           // ******************************************************************************************************
       100:  // Error state
           IF #ILx2T_Ref.ProChAccessID = #inAccessID THEN
               #ILx2T_Ref.ProChAccessID := 0;   // release access to proccessdata channel
           END_IF;
           #q_xBusy := FALSE;
           #q_xError := TRUE;
           #inState := 110;
           // ******************************************************************************************************
       110:  // finished
           IF NOT #i_xForward AND NOT #i_xBackward THEN
               #q_xError := FALSE;
               #q_xBusy := FALSE;
               #q_xCommandAborted := FALSE;
               #inState := 0;
           END_IF;
           // ******************************************************************************************************
   END_CASE;
END_FUNCTION_BLOCK

FUNCTION_BLOCK "ILx2T_Parameter_Read_Write"   // FB5, SCL
{ S7_Optimized_Access := 'TRUE' }
VERSION : 1.5
   VAR_INPUT
      i_xParameterRead : Bool;   // TRUE = Reading value continuously
      i_xParameterWrite : Bool;   // rising edge = Writing once
      i_woParameterAddress : Word;   // Parameter address (see product manual)
      i_byWriteParameterLength : Byte;   // parameter length in bytes ( 2 or 4 bytes)
      i_diWriteParameterValue : DInt;   // parameter write value
   END_VAR
   VAR_OUTPUT
      q_xReadValueValid : Bool;   // reading value is valid
      q_xWriteDone : Bool;   // writing finished without error
      q_xError : Bool;   // finished with error
      q_xBusy : Bool;   // function is active
      q_diReadParameterValue : DInt;   // reading value
   END_VAR
   VAR_IN_OUT
      ILx2T_Ref : "ILx2T_Ref";   // Axis reference structure
   END_VAR
   VAR
      inState : Int;   // internal state machine
      inAccessID : Int;   // own access ID
      inErrorState : Int;
      dwParaChErrorNo : DWord;   // parameter channe error ID
      xHelperWrite : Bool;
      xHelperRead : Bool;
      TON_Timeout : TON_TIME;
   END_VAR
BEGIN
   // *******************************************************************************
   // Init after Restart
   // *******************************************************************************
   // Check for PLC restart (1st call of this FB)
   IF #inAccessID = 0 THEN
       #ILx2T_Ref.InitAccessID := #ILx2T_Ref.InitAccessID + 1;
       #inAccessID := #ILx2T_Ref.InitAccessID;
   END_IF;

   CASE #inState OF
           // ******************************************************************************************************
       0:  // idle state
           IF #i_xParameterWrite XOR #i_xParameterRead THEN
               #xHelperWrite := #i_xParameterWrite;
               #xHelperRead := #i_xParameterRead;
               #q_xBusy := TRUE;
               #inErrorState := 0;
               #dwParaChErrorNo := 0;
               #inState := #inState + 1;
           ELSE
               #q_xWriteDone := FALSE;
               #q_xError := FALSE;
               #q_xBusy := FALSE;
               #q_xReadValueValid := FALSE;
               #q_diReadParameterValue := 0;
           END_IF;
           // ******************************************************************************************************
       1:  // Check for parameterchannel access
           IF #ILx2T_Ref.ParChAccessID = 0 OR #ILx2T_Ref.ParChAccessID = #inAccessID THEN
               #ILx2T_Ref.ParChAccessID := #inAccessID;   // grab access to parameter channel
               #inState := #inState + 1;
           END_IF;
           // ******************************************************************************************************
       2:// Prepare parameterchannel command
           #TON_Timeout(IN := FALSE,
                        PT := t#1s);
           IF #xHelperRead THEN
               #ILx2T_Ref.x_CommandReadParameter := TRUE;
               #ILx2T_Ref.udi_ModbusAddress_Read := #i_woParameterAddress;
               #inState := #inState + 1;
           ELSIF #xHelperWrite THEN
               #ILx2T_Ref.x_CommandWriteParameter := TRUE;
               #ILx2T_Ref.udi_ModbusAddress_Write := #i_woParameterAddress;
               #ILx2T_Ref.di_ParameterWriteValue := #i_diWriteParameterValue;
               #inState := #inState + 1;
           END_IF;
           // ******************************************************************************************************
       3: // Check for Parameterchannel response
           #TON_Timeout(IN := TRUE,
                        PT := t#1s);
           IF #TON_Timeout.Q THEN
               #TON_Timeout(IN := FALSE,
                            PT := t#1s);
               #q_xError := TRUE;
               #inErrorState := #inState;
               #inState := 100;
               // Read Done    
           ELSIF #xHelperRead AND #ILx2T_Ref.x_StatusReadParameter_OK AND NOT #ILx2T_Ref.x_StatusReadParameter_Error THEN
               #TON_Timeout(IN := FALSE,
                            PT := t#1s);
               #q_diReadParameterValue := #ILx2T_Ref.di_ParameterReadValue;
               #q_xReadValueValid := TRUE;
               #ILx2T_Ref.x_CommandReadParameter := FALSE;
               #ILx2T_Ref.x_StatusReadParameter_OK := FALSE;
               #ILx2T_Ref.udi_ModbusAddress_Read := 0;
               #inState := #inState + 1;
               // Write Done    
           ELSIF #xHelperWrite AND #ILx2T_Ref.x_Status_WriteParameter_OK AND NOT #ILx2T_Ref.x_Status_WriteParameter_Error THEN
               #TON_Timeout(IN := FALSE,
                            PT := t#1s);
               #ILx2T_Ref.di_ParameterWriteValue := 0;
               #q_xWriteDone := TRUE;
               #ILx2T_Ref.x_CommandWriteParameter := FALSE;
               #ILx2T_Ref.x_Status_WriteParameter_OK := FALSE;
               #ILx2T_Ref.udi_ModbusAddress_Write := 0;
               #inState := #inState + 1;
               // Error response Reading
           ELSIF #ILx2T_Ref.x_StatusReadParameter_Error THEN
               #ILx2T_Ref.x_CommandReadParameter := FALSE;
               #ILx2T_Ref.x_StatusReadParameter_Error := FALSE;
               #ILx2T_Ref.udi_ModbusAddress_Read := 0;
               #TON_Timeout(IN := FALSE,
                            PT := t#1s);
               #inErrorState := #inState;
               #inState := 100;
               // Error response Writing
           ELSIF #ILx2T_Ref.x_Status_WriteParameter_Error THEN
               #ILx2T_Ref.x_CommandWriteParameter := FALSE;
               #ILx2T_Ref.x_Status_WriteParameter_Error := FALSE;
               #ILx2T_Ref.udi_ModbusAddress_Write := 0;
               #TON_Timeout(IN := FALSE,
                            PT := t#1s);
               #inErrorState := #inState;
               #inState := 100;
           END_IF;
           // ******************************************************************************************************
       4:  // Check for Parameterchannel in idle state
           #TON_Timeout(IN := TRUE,
                        PT := t#1s);
           IF #TON_Timeout.Q THEN
               #TON_Timeout(IN := FALSE,
                            PT := t#1s);
               #q_xError := TRUE;
               #inErrorState := #inState;
               #inState := 100;
           ELSIF NOT #ILx2T_Ref.x_StatusReadParameter_OK AND NOT #ILx2T_Ref.x_StatusReadParameter_Error
               AND NOT #ILx2T_Ref.x_Status_WriteParameter_OK AND NOT #ILx2T_Ref.x_Status_WriteParameter_Error THEN
               #ILx2T_Ref.ParChAccessID := 0;   // grab access to parameter channel
               #TON_Timeout(IN := FALSE,
                            PT := t#1s);
               IF #xHelperWrite THEN
                   #q_xBusy := FALSE;
                   #inState := 110;
               ELSE
                   #inState := 0;
               END_IF;
           END_IF;
       100:  // Error state
           IF #ILx2T_Ref.ParChAccessID = #inAccessID THEN
               #ILx2T_Ref.ParChAccessID := 0;   // release access to proccessdata channel
           END_IF;
           #q_xBusy := FALSE;
           #q_xError := TRUE;
           #inState := 110;
           // ******************************************************************************************************
       110:  // finished
           IF NOT #i_xParameterWrite AND NOT #i_xParameterRead THEN
               #q_xWriteDone := FALSE;
               #q_xError := FALSE;
               #q_xBusy := FALSE;
               #q_xReadValueValid := FALSE;
               #q_diReadParameterValue := 0;
               #inState := 0;
           END_IF;
           // ******************************************************************************************************
   END_CASE;
END_FUNCTION_BLOCK

FUNCTION_BLOCK "ILx2T_ProfilePosition"   // FB6, SCL
{ S7_Optimized_Access := 'TRUE' }
VERSION : 1.5
   VAR_INPUT
      i_xExecute : Bool;   // rising edge starts a new movement
      i_xAbort : Bool;   // abort active movement
      i_inPTP_Type : Int;   // 1=absolute / 2=additive / 3=relative
      i_diTargetPosition : DInt;   // Target position value
      i_inTargetVelocity : Int;   // Target velocity value
   END_VAR
   VAR_OUTPUT
      q_xDone : Bool;   // Target position reached
      q_xError : Bool;   // finished with error
      q_xCommandAborted : Bool;   // function aborted
      q_xBusy : Bool;   // function is active
   END_VAR
   VAR_IN_OUT
      ILx2T_Ref : "ILx2T_Ref";   // Axis reference structure
   END_VAR
   VAR
      inState : Int;   // internal state machine
      inAccessID : Int;   // own access ID
      inHelperState : Int;
      inErrorState : Int;
      woInternalErrorID : Word;   // internal FB error ID
      xModeToggleHelper : Bool;
      xHelperExecute : Bool;
      inHelperTargetVelocity : Int;
      TON_Timeout : TON_TIME;
   END_VAR
BEGIN
   // *******************************************************************************
   // Init after Restart
   // *******************************************************************************
   // Check for PLC restart (1st call of this FB)
   IF #inAccessID = 0 THEN
       #ILx2T_Ref.InitAccessID := #ILx2T_Ref.InitAccessID + 1;
       #inAccessID := #ILx2T_Ref.InitAccessID;
   END_IF;

   CASE #inState OF
           // ******************************************************************************************************
       0:  // idle state
           IF #i_xExecute THEN
               #q_xBusy := TRUE;
               #inErrorState := 0;
               #inState := #inState + 1;
           ELSE
               #q_xDone := FALSE;
               #q_xError := FALSE;
               #q_xBusy := FALSE;
               #q_xCommandAborted := FALSE;
           END_IF;
           // ******************************************************************************************************
       1:  // Check for drive state and access ID
           IF NOT #ILx2T_Ref.stDriveStatus.x_End AND #ILx2T_Ref.by_OP_ModeAct <> 3 THEN  // A318 operating mode active
               #q_xError := TRUE;
               #woInternalErrorID := 16#A318;
               #inErrorState := #inState;
               #inState := 100;
           ELSIF (#ILx2T_Ref.i_woDriveStatus AND 16#F) = 6 THEN
               #inState := #inState + 1;
           ELSE
               #q_xError := TRUE;
               #inErrorState := #inState;
               #inState := 100;
           END_IF;
           // ******************************************************************************************************
       2: // Start Movement via Processchannel
           //   i_inPTP_Type 1 = Mode 03 hex = move absolute (RefA32 = target velocity / RefB32 = target position)
           //   i_inPTP_Type 2 = Mode 13 hex = move additive (RefA32 = target velocity / RefB32 = target position)
           //   i_inPTP_Type 3 = Mode 23 hex = move relative (RefA32 = target velocity / RefB32 = target position)
           #ILx2T_Ref.q_dw_refA_16 := INT_TO_WORD(#i_inTargetVelocity);
           #inHelperTargetVelocity := #i_inTargetVelocity;
           #ILx2T_Ref.q_dw_refB_32 := DINT_TO_DWORD(#i_diTargetPosition);
           #xHelperExecute := FALSE;
           CASE #i_inPTP_Type OF
               1: // Move absolute
                   #ILx2T_Ref.q_wo_dmControl := #ILx2T_Ref.q_wo_dmControl AND 16#FF80;
                   #ILx2T_Ref.q_wo_dmControl := #ILx2T_Ref.q_wo_dmControl OR 16#0003;
                   #inState := #inState + 1;
               2: // Move additive
                   #ILx2T_Ref.q_wo_dmControl := #ILx2T_Ref.q_wo_dmControl AND 16#FF80;
                   #ILx2T_Ref.q_wo_dmControl := #ILx2T_Ref.q_wo_dmControl OR 16#0013;
                   #inState := #inState + 1;
               3: // Move relative
                   #ILx2T_Ref.q_wo_dmControl := #ILx2T_Ref.q_wo_dmControl AND 16#FF80;
                   #ILx2T_Ref.q_wo_dmControl := #ILx2T_Ref.q_wo_dmControl OR 16#0023;
                   #inState := #inState + 1;
               ELSE
                   #inErrorState := #inState;
                   #inState := 100;
           END_CASE;

           // ******************************************************************************************************
       3: // ModeToggle 
           IF NOT #i_xExecute THEN
               #xHelperExecute := TRUE;
           END_IF;
           #xModeToggleHelper := NOT #ILx2T_Ref.st_ModeStatus.ModeToggle;  // save toggle bit 
           IF NOT #xModeToggleHelper THEN
               #ILx2T_Ref.q_wo_dmControl := #ILx2T_Ref.q_wo_dmControl AND 16#FF7F;
           ELSE
               #ILx2T_Ref.q_wo_dmControl := #ILx2T_Ref.q_wo_dmControl OR 16#0080;
           END_IF;
           #inState := #inState + 1;
           // ******************************************************************************************************
       4: // Check for mode toggle and number of operating mode OK
           IF NOT #i_xExecute THEN
               #xHelperExecute := TRUE;
           END_IF;
           IF NOT (#xModeToggleHelper XOR #ILx2T_Ref.st_ModeStatus.ModeToggle) AND (#ILx2T_Ref.by_OP_ModeAct = 16#0003) THEN                            // Check operating mode number
               #TON_Timeout(IN := FALSE,
                            PT := t#1s);
               #inState := #inState + 1;  // Command OK
           ELSE
               // TIMEOUT ERROR
               #TON_Timeout(IN := TRUE,
                            PT := t#1s);
               IF #TON_Timeout.Q THEN
                   #TON_Timeout(IN := FALSE,
                                PT := t#1s);
                   #q_xError := TRUE;
                   #inErrorState := #inState;
                   #inState := 100;
               END_IF;
           END_IF;
           // ******************************************************************************************************
       5: // Check operating mode
           IF NOT #i_xExecute THEN
               #xHelperExecute := TRUE;
           END_IF;
           // Mode OK -> Check drive status (x_Add, x_End and x_Error)
           IF #ILx2T_Ref.stDriveStatus.x_Add AND #ILx2T_Ref.stDriveStatus.x_End AND NOT #ILx2T_Ref.stDriveStatus.x_Err THEN  // finished without Error     
               #q_xBusy := FALSE;
               #q_xDone := TRUE;
               #inState := 110;
           ELSIF #ILx2T_Ref.stDriveStatus.x_End AND #ILx2T_Ref.stDriveStatus.x_Err THEN  // finished with Error     
               #inErrorState := #inState;
               #inState := 100;
           ELSIF #ILx2T_Ref.by_OP_ModeAct <> 16#0003 THEN   // check for correct operating mode number
               #q_xCommandAborted := TRUE;
               #q_xBusy := FALSE;
               #q_xDone := FALSE;
               #inState := 110;
           ELSIF #i_xExecute AND #xHelperExecute THEN
               #inState := 2;
           ELSIF #i_xAbort THEN
               #ILx2T_Ref.x_QuickStopInt := TRUE;
               #inState := #inState + 1;
           // Velocity can be changed during movement (only move absolute)
           ELSIF #i_inPTP_Type = 1 THEN
               IF #inHelperTargetVelocity <> #i_inTargetVelocity THEN
                   #inState := 2;
               END_IF;
           END_IF;
       6:
           IF #ILx2T_Ref.stDriveStatus.x_End AND (#ILx2T_Ref.i_woDriveStatus AND 16#F) >= 7 THEN  // Check for STANDSTILL
               #ILx2T_Ref.x_QuickStopInt := FALSE;
               #ILx2T_Ref.x_FaultResetInt := TRUE;
               #TON_Timeout(IN := TRUE,
                            PT := t#1s);
               IF #TON_Timeout.Q THEN
                   #TON_Timeout(IN := FALSE,
                                PT := t#1s);
                   #ILx2T_Ref.x_FaultResetInt := FALSE;
                   #q_xError := TRUE;
                   #inErrorState := #inState;
                   #inState := 100;
               END_IF;
           ELSIF #ILx2T_Ref.stDriveStatus.x_End AND (#ILx2T_Ref.i_woDriveStatus AND 16#F) < 7 THEN  // Check for STANDSTILL
               #ILx2T_Ref.x_QuickStopInt := FALSE;
               #ILx2T_Ref.x_FaultResetInt := FALSE;
               #q_xCommandAborted := TRUE;
               #q_xBusy := FALSE;
               #q_xDone := FALSE;
               #inState := 110;
           END_IF;

           // ******************************************************************************************************
       100:  // Error state
           #q_xBusy := FALSE;
           #q_xError := TRUE;
           #inState := 110;
           // ******************************************************************************************************
       110:  // finished
           IF NOT #i_xExecute AND NOT #i_xAbort THEN
               #q_xDone := FALSE;
               #q_xError := FALSE;
               #q_xBusy := FALSE;
               #q_xCommandAborted := FALSE;
               #inState := 0;
           END_IF;
           // ******************************************************************************************************
   END_CASE;
END_FUNCTION_BLOCK

FUNCTION_BLOCK "ILx2T_ProfileVelocity"   // FB8, SCL
{ S7_Optimized_Access := 'TRUE' }
VERSION : 1.5
   VAR_INPUT
      i_xExecute : Bool;   // Start movement
      i_xAbort : Bool;   // Abort current movement
      i_inTargetVelocity : Int;   // Target speed
   END_VAR
   VAR_OUTPUT
      q_xTargetVelocityReached : Bool;   // Target velocity reached
      q_xError : Bool;   // FB finished with error
      q_xCommandAborted : Bool;   // FB aborted
      q_xBusy : Bool;   // function block is busy
   END_VAR
   VAR_IN_OUT
      ILx2T_Ref : "ILx2T_Ref";   // Axis reference structure
   END_VAR
   VAR
      inState : Int;   // internal state machine
      inAccessID : Int;   // own access ID
      inHelperState : Int;
      inErrorState : Int;
      woInternalErrorID : Word;   // internal FB error ID
      xModeToggleHelper : Bool;
      inTargetVelocityHelper : Int;
      TON_Timeout : TON_TIME;
   END_VAR
BEGIN
   // *******************************************************************************
   // Init after Restart
   // *******************************************************************************
   // Check for PLC restart (1st call of this FB)
   IF #inAccessID = 0 THEN
       #ILx2T_Ref.InitAccessID := #ILx2T_Ref.InitAccessID + 1;
       #inAccessID := #ILx2T_Ref.InitAccessID;
   END_IF;

   CASE #inState OF
           // ******************************************************************************************************
       0:  // idle state
           IF #i_xExecute THEN
               #q_xBusy := TRUE;
               #inErrorState := 0;
               #inState := #inState + 1;
           ELSE
               #q_xTargetVelocityReached := FALSE;
               #q_xError := FALSE;
               #q_xBusy := FALSE;
               #q_xCommandAborted := FALSE;
           END_IF;
           // ******************************************************************************************************
       1:  // Check for drive state and access ID
           IF NOT #ILx2T_Ref.stDriveStatus.x_End AND #ILx2T_Ref.by_OP_ModeAct <> 4 THEN  // A318 operating mode active
               #q_xError := TRUE;
               #woInternalErrorID := 16#A318;
               #inErrorState := #inState;
               #inState := 100;
           ELSIF (#ILx2T_Ref.i_woDriveStatus AND 16#F) = 6 THEN
               #inState := #inState + 1;
           ELSE
               #q_xError := TRUE;
               #inErrorState := #inState;
               #inState := 100;
           END_IF;
           // ******************************************************************************************************

           // ******************************************************************************************************
       2: // Start Movement via Processchannel
           // Mode 04 hex = Profile Velocity (RefA32 = target velocity / RefB32 = reserved)
           #ILx2T_Ref.q_dw_refB_32 := 0;
           #ILx2T_Ref.q_dw_refA_16 := INT_TO_WORD(#i_inTargetVelocity);
           #inTargetVelocityHelper := #i_inTargetVelocity;
           #ILx2T_Ref.q_wo_dmControl := #ILx2T_Ref.q_wo_dmControl AND 16#FF80;
           #ILx2T_Ref.q_wo_dmControl := #ILx2T_Ref.q_wo_dmControl OR 16#0004;
           #inState := #inState + 1;
           // ******************************************************************************************************
       3: // Mode Toggle
           #xModeToggleHelper := NOT #ILx2T_Ref.st_ModeStatus.ModeToggle;   // save toggle bit 
           IF NOT #xModeToggleHelper THEN
               #ILx2T_Ref.q_wo_dmControl := #ILx2T_Ref.q_wo_dmControl AND 16#FF7F;
           ELSE
               #ILx2T_Ref.q_wo_dmControl := #ILx2T_Ref.q_wo_dmControl OR 16#0080;
           END_IF;
           #inState := #inState + 1;
           // ******************************************************************************************************
       4: // Check for mode response OK
           // Check for mode toggle and number of operating mode OK
           IF NOT (#xModeToggleHelper XOR #ILx2T_Ref.st_ModeStatus.ModeToggle) AND (#ILx2T_Ref.by_OP_ModeAct = 16#0004) THEN                            // Check operating mode number
               #TON_Timeout(IN := FALSE,
                            PT := t#1s);
               #inState := #inState + 1;
           ELSE
               // TIMEOUT ERROR
               #TON_Timeout(IN := TRUE,
                            PT := t#1s);
               IF #TON_Timeout.Q THEN
                   #TON_Timeout(IN := FALSE,
                                PT := t#1s);
                   #q_xError := TRUE;
                   #inErrorState := #inState;
                   #inState := 100;
               END_IF;
           END_IF;
           // ******************************************************************************************************
       5: // Check operating mode
           // Check for target reached (Drive status x_Add)
           IF (#ILx2T_Ref.i_woDriveStatus AND 16#2000) = 16#2000 THEN  // x_Add = Target vel reached     
               #q_xTargetVelocityReached := TRUE;
           ELSE
               #q_xTargetVelocityReached := FALSE;
           END_IF;
           // x_Error
           IF (#ILx2T_Ref.i_woDriveStatus AND 16#8000) = 16#8000 THEN  // error     
               #inErrorState := #inState;
               #inState := 100;
           // Monitoring of actual operating mode
           ELSIF (#ILx2T_Ref.by_OP_ModeAct <> 16#0004) THEN
               #q_xCommandAborted := TRUE;
               #q_xBusy := FALSE;
               #q_xTargetVelocityReached := FALSE;
               #inState := 110;
           // Check for new target velocity value !
           ELSIF #inTargetVelocityHelper <> #i_inTargetVelocity THEN
               #inState := 2;
           // Check for ABORT command
           ELSIF #i_xAbort THEN
               #ILx2T_Ref.x_QuickStopInt := TRUE;
               #inState := #inState + 1;
           END_IF;
       6:
           #TON_Timeout(IN := TRUE,
                        PT := t#10s);
           IF #TON_Timeout.Q THEN
               #TON_Timeout(IN := FALSE,
                            PT := t#1s);
               #ILx2T_Ref.x_QuickStopInt := FALSE;
               #ILx2T_Ref.x_FaultResetInt := FALSE;
               #q_xError := TRUE;
               #inErrorState := #inState;
               #inState := 100;
           ELSIF #ILx2T_Ref.stDriveStatus.x_End AND (#ILx2T_Ref.i_woDriveStatus AND 16#F) >= 7 THEN  // Check for STANDSTILL
               #ILx2T_Ref.x_QuickStopInt := FALSE;
               #ILx2T_Ref.x_FaultResetInt := TRUE;
           ELSIF #ILx2T_Ref.stDriveStatus.x_End AND (#ILx2T_Ref.i_woDriveStatus AND 16#F) < 7 THEN  // Check for STANDSTILL
               #TON_Timeout(IN := FALSE,
                            PT := t#1s);
               #ILx2T_Ref.x_QuickStopInt := FALSE;
               #ILx2T_Ref.x_FaultResetInt := FALSE;
               #q_xCommandAborted := TRUE;
               #q_xBusy := FALSE;
               #q_xTargetVelocityReached := FALSE;
               #inState := 110;
           END_IF;

           // ******************************************************************************************************
       100:  // Error state
           #q_xBusy := FALSE;
           #q_xError := TRUE;
           #inState := 110;
           // ******************************************************************************************************
       110:  // finished
           IF NOT #i_xExecute AND NOT #i_xAbort THEN
               #q_xTargetVelocityReached := FALSE;
               #q_xError := FALSE;
               #q_xBusy := FALSE;
               #q_xCommandAborted := FALSE;
               #inState := 0;
           END_IF;
           // ******************************************************************************************************
   END_CASE;
END_FUNCTION_BLOCK

FUNCTION_BLOCK "ILx2_ModbusTCP_Data_1500"   // FB10, SCL
{ S7_Optimized_Access := 'FALSE' }
VERSION : 1.5
   VAR_INPUT
      CONNECT_ID_1 : Conn_Ouc := 1;   // unique connection ID DPL Read
      CONNECT_ID_2 : Conn_Ouc := 2;   // unique connection ID DPL Write
      CONNECT_ID_3 : Conn_Ouc := 3;   // unique connection ID Parameter read
      CONNECT_ID_4 : Conn_Ouc := 4;   // unique connection ID Parameter write
      IP_OCTET_1 : USInt := 192;
      IP_OCTET_2 : USInt := 168;
      IP_OCTET_3 : USInt;
      IP_OCTET_4 : USInt;
      inNodeGuardTime : UInt := 1000;   // Modbus Node Guard Time (Object 6544 Range 0..10000 ms)
   END_VAR
   VAR_OUTPUT
      Com_OK : Bool;   // Communication OK
      Error : Bool;   // Communication error
      ErrorCode : Word;   // MB_CLIENT - error code
   END_VAR
   VAR_IN_OUT
      ILx2T_Ref : "ILx2T_Ref";
   END_VAR
   VAR
      ReadData_DPL : Array[0..7] of Byte;   // Read Data Drive Profile Lexium
      WriteData_DPL : Array[0..7] of Byte;   // Write Data Drive Profile Lexium
      ParaRead_Value : DInt;   // Parameter Read Data
      ParaWrite_Value : DInt;   // Parameter Write Data
      iState_Read_DPL : Int;
      iState_Write_DPL : Int;
      iState_Read_Para : Int;
      iState_Write_Para : Int;
      MB_CLIENT_Instance_DPL_Read : MB_CLIENT;
      MB_CLIENT_Instance_DPL_Write : MB_CLIENT;
      MB_CLIENT_Instance_ParaRead : MB_CLIENT;
      MB_CLIENT_Instance_ParaWrite : MB_CLIENT;
      stCONNECT_DPL_Read : TCON_IP_v4;
      stCONNECT_DPL_Write : TCON_IP_v4;
      stCONNECT_Parameter_Read : TCON_IP_v4;
      stCONNECT_Parameter_Write : TCON_IP_v4;
      Index : Int;
      inIndex : Int;
      xNodeGuardInitOK : Bool;
      xErrorReadDPL : Bool;
      xErrorWriteDPL : Bool;
      xErrorReadParameter : Bool;
      xErrorWriteParameter : Bool;
      diErrorCounter_DPL_Read : DInt;
      diErrorCounter_DPL_Write : DInt;
      diErrorCounter_Para_Read : DInt;
      diErrorCounter_Para_Write : DInt;
      woReadDPL_ErrorID : Word;
      woWriteDPL_ErrorID : Word;
      woReadParameter_ErrorID : Word;
      woWriteParameter_ErrorID : Word;
      iStateTimeReadDPL : Int;
      iStateTimeWriteDPL : Int;
      T_ReadDPL : TON_TIME;
      t_ReadDPL_Min : Time := t#5m;
      t_ReadDPL_Act : Time;
      t_ReadDPL_Max : Time;
      T_WriteDPL : TON_TIME;
      t_WriteDPL_Min : Time := t#5m;
      t_WriteDPL_Act : Time;
      t_WriteDPL_Max : Time;
      MB_CLIENT_Instance : MB_CLIENT;
   END_VAR
BEGIN
   // THIS FB uses ModbusTCP 5.0 - 04.02.2019
   // OpenUserCommunication must be set to Version 5.1 - 04.02.2019
   // 23.07.2018 - Using 4 connections to increase the performance of the data exchange
   // ***************************************************************************************
   // S7-1x00 - MB_Client Version 5.0
   // PLC IP address 10.209.177.xxx
   // Modbus slave IP Address 10.209.177.xxx
   // ***************************************************************************************
   // Read DPL Data OF 4 WORDS from slave
   // ***************************************************************************************
   #stCONNECT_DPL_Read.ActiveEstablished := TRUE;
   #stCONNECT_DPL_Read.ConnectionType := 11;    // TCP
   #stCONNECT_DPL_Read.ID := #CONNECT_ID_1;
   #stCONNECT_DPL_Read.InterfaceId := 64;    // PROFINET Network
   #stCONNECT_DPL_Read.LocalPort := 0;
   #stCONNECT_DPL_Read.RemotePort := 502;   // 502 See TIA ONLINE HELP
   #stCONNECT_DPL_Read.RemoteAddress.ADDR[1] := #IP_OCTET_1;
   #stCONNECT_DPL_Read.RemoteAddress.ADDR[2] := #IP_OCTET_2;
   #stCONNECT_DPL_Read.RemoteAddress.ADDR[3] := #IP_OCTET_3;
   #stCONNECT_DPL_Read.RemoteAddress.ADDR[4] := #IP_OCTET_4;
   CASE #iState_Read_DPL OF
       0:  // DISCONNECT
           #MB_CLIENT_Instance_DPL_Read(REQ := FALSE,
                                        DISCONNECT := TRUE,
                                        MB_MODE := 0,
                                        MB_DATA_ADDR := 400001 + 6926,
                                        MB_DATA_LEN := 4,
                                        MB_DATA_PTR := #ReadData_DPL,
                                        CONNECT := #stCONNECT_DPL_Read);
           #iState_Read_DPL := #iState_Read_DPL + 1;
       1:  // CONNECT  
           #MB_CLIENT_Instance_DPL_Read(REQ := false,
                                        DISCONNECT := FALSE,
                                        MB_MODE := 0,
                                        MB_DATA_ADDR := 400001 + 6926,
                                        MB_DATA_LEN := 4,
                                        MB_DATA_PTR := #ReadData_DPL,
                                        CONNECT := #stCONNECT_DPL_Read);
           IF #MB_CLIENT_Instance_DPL_Read.Connected AND NOT #MB_CLIENT_Instance_DPL_Read.BUSY THEN
               IF NOT #xNodeGuardInitOK THEN
                   #iState_Read_DPL := 200;
               ELSE
                   #iState_Read_DPL := #iState_Read_DPL + 1;
               END_IF;
           ELSIF #MB_CLIENT_Instance_DPL_Read.ERROR THEN
               #woReadDPL_ErrorID := #MB_CLIENT_Instance_DPL_Read.STATUS;
               #iState_Read_DPL := #iState_Read_DPL + 100;
           END_IF;
       2:  // Check for DONE AND NOT BUSY
           #MB_CLIENT_Instance_DPL_Read(REQ := TRUE,
                                        DISCONNECT := FALSE,
                                        MB_MODE := 0,
                                        MB_DATA_ADDR := 400001 + 6926,
                                        MB_DATA_LEN := 4,
                                        MB_DATA_PTR := #ReadData_DPL,
                                        CONNECT := #stCONNECT_DPL_Read);
           IF #MB_CLIENT_Instance_DPL_Read.DONE AND NOT #MB_CLIENT_Instance_DPL_Read.BUSY THEN
               #xErrorReadDPL := FALSE;
               #woReadDPL_ErrorID := 0;
               FOR #Index := 0 TO 7 DO
                   #ILx2T_Ref.arInputData[#Index] := #ReadData_DPL[#Index];
               END_FOR;
           ELSIF #MB_CLIENT_Instance_DPL_Read.ERROR THEN
               #woReadDPL_ErrorID := #MB_CLIENT_Instance_DPL_Read.STATUS;
               FOR #Index := 0 TO 7 DO
                   #ILx2T_Ref.arInputData[#Index] := 0;
               END_FOR;
               #iState_Read_DPL := #iState_Read_DPL + 100;
           END_IF;
       100..120:  // Error state
           #xErrorReadDPL := TRUE;
           #diErrorCounter_DPL_Read := #diErrorCounter_DPL_Read + 1;
           #MB_CLIENT_Instance_DPL_Read(REQ := FALSE,
                                        DISCONNECT := TRUE,
                                        MB_MODE := 0,
                                        MB_DATA_ADDR := 400001 + 6926,
                                        MB_DATA_LEN := 4,
                                        MB_DATA_PTR := #ReadData_DPL,
                                        CONNECT := #stCONNECT_DPL_Read);
           #iState_Read_DPL := 0;

           // **********************************************************************************************************
           // ***** Set Modbus Nodeguar time after communication is established once ***********************************
           // **********************************************************************************************************
       200:  // CONNECT  
           #ParaWrite_Value := #inNodeGuardTime;
           #MB_CLIENT_Instance_DPL_Read(REQ := FALSE,
                                        DISCONNECT := FALSE,
                                        MB_MODE := 1,
                                        MB_DATA_ADDR := 400001 + 5644,
                                        MB_DATA_LEN := 2,
                                        MB_DATA_PTR := #ParaWrite_Value,
                                        CONNECT := #stCONNECT_DPL_Read);
           IF #MB_CLIENT_Instance_DPL_Read.Connected AND NOT #MB_CLIENT_Instance_DPL_Read.BUSY THEN
               #woReadDPL_ErrorID := 0;
               #iState_Read_DPL := #iState_Read_DPL + 1;
           ELSIF #MB_CLIENT_Instance_DPL_Read.ERROR THEN
               #woReadDPL_ErrorID := #MB_CLIENT_Instance_DPL_Read.STATUS;
               #iState_Read_DPL := 119;
           END_IF;
       201:  // Write Parameter
           #ParaWrite_Value := #inNodeGuardTime;
           #MB_CLIENT_Instance_DPL_Read(REQ := TRUE,
                                        DISCONNECT := FALSE,
                                        MB_MODE := 1,
                                        MB_DATA_ADDR := 400001 + 5644,
                                        MB_DATA_LEN := 2,
                                        MB_DATA_PTR := #ParaWrite_Value,
                                        CONNECT := #stCONNECT_DPL_Read);
           IF #MB_CLIENT_Instance_DPL_Read.DONE AND NOT #MB_CLIENT_Instance_DPL_Read.BUSY THEN
               #woReadDPL_ErrorID := 0;
               #MB_CLIENT_Instance_DPL_Read(REQ := FALSE,
                                            DISCONNECT := FALSE,
                                            MB_MODE := 1,
                                            MB_DATA_ADDR := 400001 + 5644,
                                            MB_DATA_LEN := 2,
                                            MB_DATA_PTR := #ParaWrite_Value,
                                            CONNECT := #stCONNECT_DPL_Read);
               #xNodeGuardInitOK := TRUE;
               #iState_Read_DPL := 0;
           ELSIF #MB_CLIENT_Instance_DPL_Read.ERROR THEN
               #woReadDPL_ErrorID := #MB_CLIENT_Instance_DPL_Read.STATUS;
               #iState_Read_DPL := 120;
           END_IF;